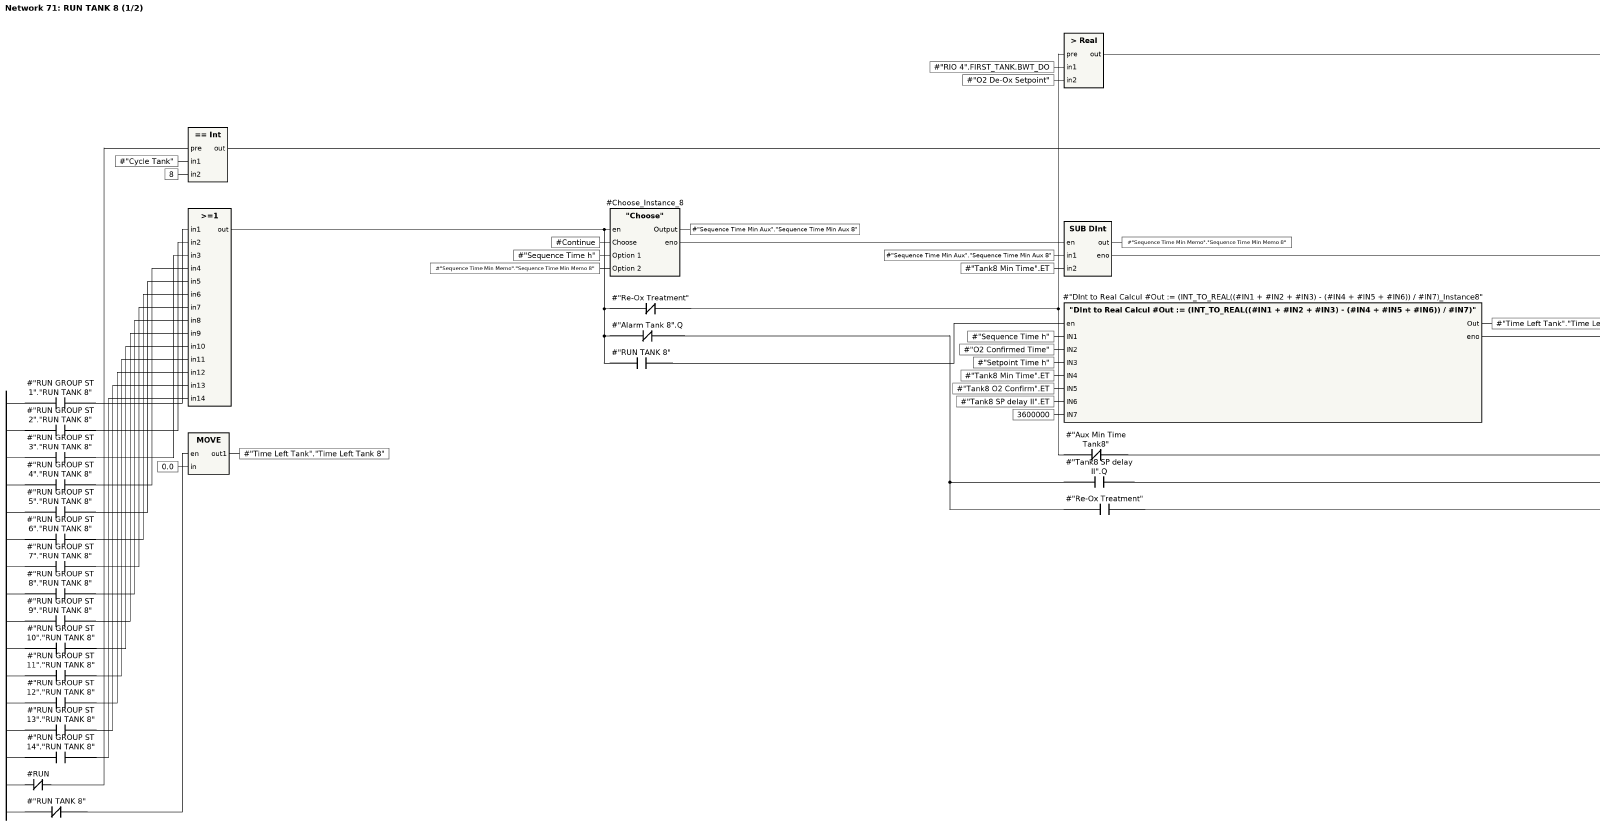
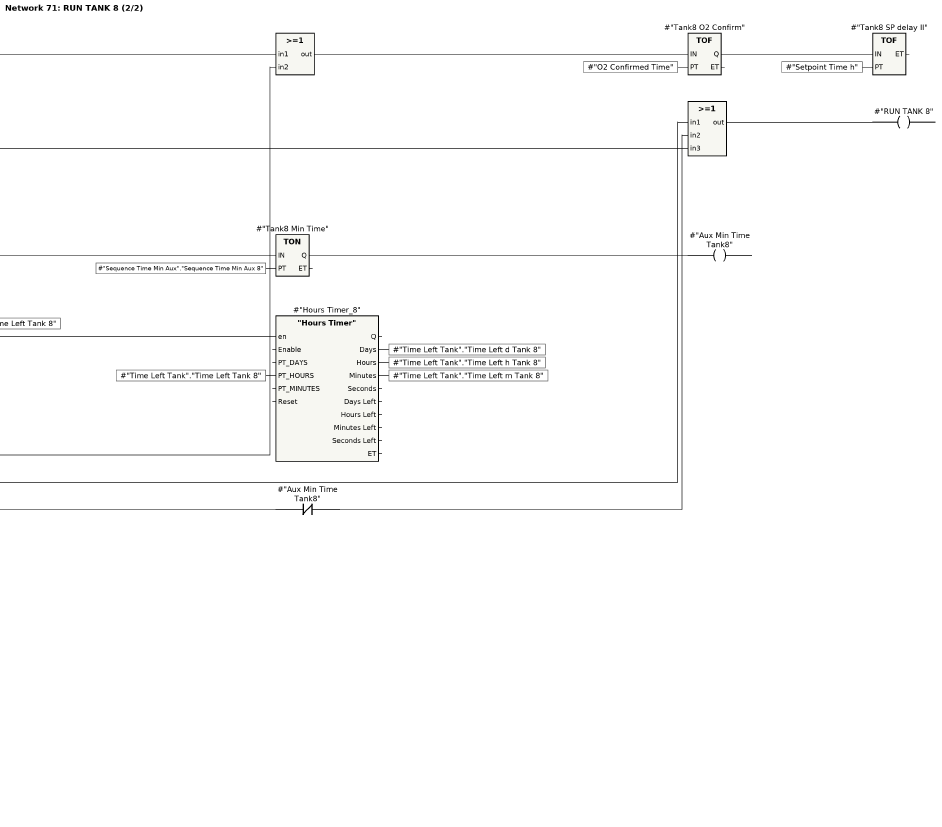
   #_w1 := #"RUN GROUP ST 1"."RUN TANK 8" OR #"RUN GROUP ST 2"."RUN TANK 8" OR #"RUN GROUP ST 3"."RUN TANK 8" OR #"RUN GROUP ST 4"."RUN TANK 8" OR #"RUN GROUP ST 5"."RUN TANK 8" OR #"RUN GROUP ST 6"."RUN TANK 8" OR #"RUN GROUP ST 7"."RUN TANK 8" OR #"RUN GROUP ST 8"."RUN TANK 8" OR #"RUN GROUP ST 9"."RUN TANK 8" OR #"RUN GROUP ST 10"."RUN TANK 8" OR #"RUN GROUP ST 11"."RUN TANK 8" OR #"RUN GROUP ST 12"."RUN TANK 8" OR #"RUN GROUP ST 13"."RUN TANK 8" OR #"RUN GROUP ST 14"."RUN TANK 8";
   #Choose_Instance_8(EN := #_w1,   // "Choose"
                      Choose := #Continue,
                      "Option 1" := #"Sequence Time h",
                      "Option 2" := #"Sequence Time Min Memo"."Sequence Time Min Memo 8",
                      Output => #"Sequence Time Min Aux"."Sequence Time Min Aux 8",
                      ENO => #_w2);
   IF #_w2 THEN
       #"Sequence Time Min Memo"."Sequence Time Min Memo 8" := #"Sequence Time Min Aux"."Sequence Time Min Aux 8" - #"Tank8 Min Time".ET;   // Memory of remained time for use to continue
   END_IF;
   #"Tank8 Min Time"(IN := #_w2, PT := #"Sequence Time Min Aux"."Sequence Time Min Aux 8");   // TON
   #"Aux Min Time Tank8" := #"Tank8 Min Time".Q;
   #"Tank8 O2 Confirm"(IN := #_w1 AND NOT #"Re-Ox Treatment" AND ((#"RIO 4".FIRST_TANK.BWT_DO > #"O2 De-Ox Setpoint") OR NOT #"Aux Min Time Tank8"),   // TOF
                       PT := #"O2 Confirmed Time");
   #"Tank8 SP delay II"(IN := #"Tank8 O2 Confirm".Q, PT := #"Setpoint Time h");   // TOF
   #"DInt to Real Calcul #Out := (INT_TO_REAL((#IN1 + #IN2 + #IN3) - (#IN4 + #IN5 + #IN6)) / #IN7)_Instance8"(EN := #_w1 AND #"RUN TANK 8",   // "DInt to Real Calcul #Out := (INT_TO_REAL((#IN1 + #IN2 + #IN3) - (#IN4 + #IN5 + #IN6)) / #IN7)"
                           IN1 := #"Sequence Time h",
                           IN2 := #"O2 Confirmed Time",
                           IN3 := #"Setpoint Time h",
                           IN4 := #"Tank8 Min Time".ET,
                           IN5 := #"Tank8 O2 Confirm".ET,
                           IN6 := #"Tank8 SP delay II".ET,
                           IN7 := 3600000,
                           Out => #"Time Left Tank"."Time Left Tank 8",
                           ENO => #_w3);
   IF #_w3 THEN
       #"Hours Timer_8"(PT_HOURS := #"Time Left Tank"."Time Left Tank 8",   // "Hours Timer"
                        Days => #"Time Left Tank"."Time Left d Tank 8",
                        Hours => #"Time Left Tank"."Time Left h Tank 8",
                        Minutes => #"Time Left Tank"."Time Left m Tank 8");
   END_IF;
   #"RUN TANK 8" := (#_w1 AND NOT #"Alarm Tank 8".Q AND (#"Tank8 SP delay II".Q OR (#"Re-Ox Treatment" AND NOT #"Aux Min Time Tank8"))) OR (NOT #RUN AND (#"Cycle Tank" = 8));
   IF NOT #"RUN TANK 8" THEN #"Time Left Tank"."Time Left Tank 8" := 0.0; END_IF;
END_REGION

REGION Network 72: RUN TANK 9
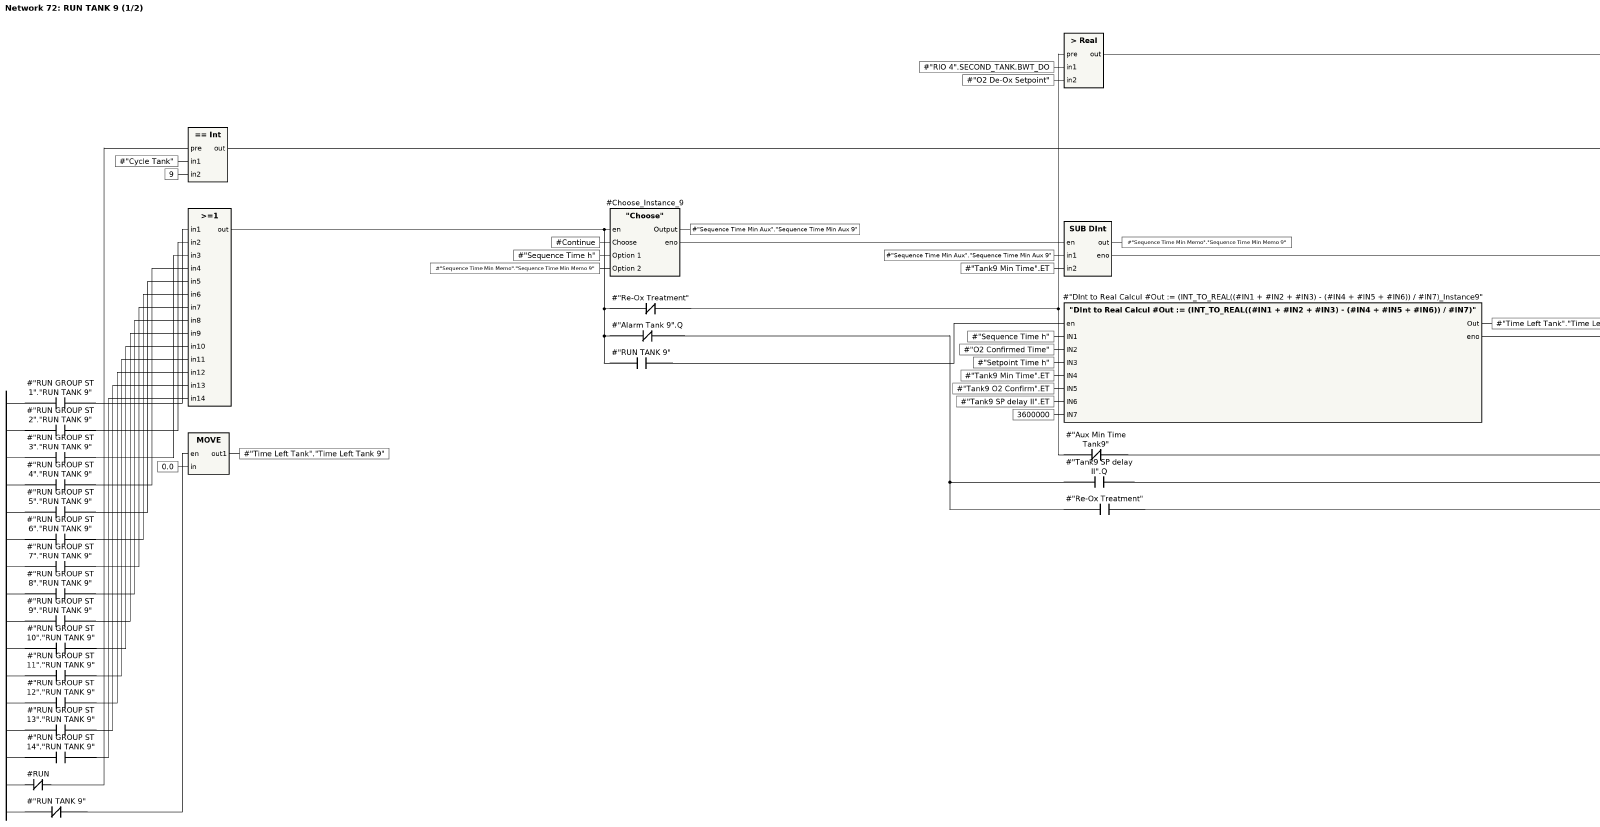
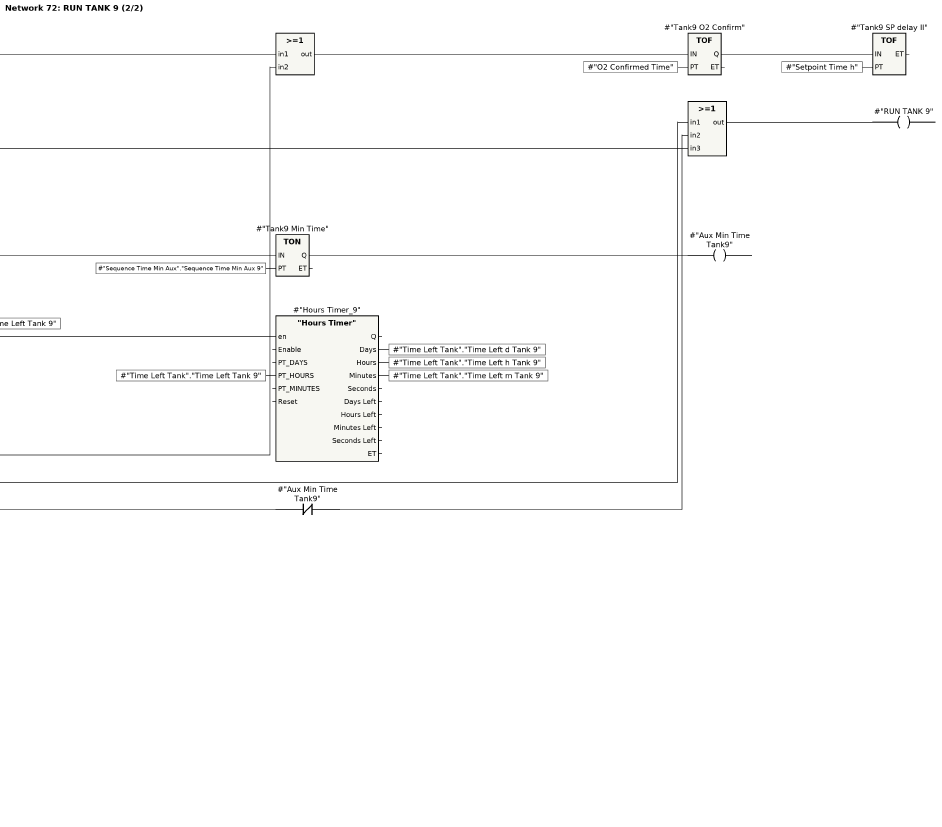
   #_w1 := #"RUN GROUP ST 1"."RUN TANK 9" OR #"RUN GROUP ST 2"."RUN TANK 9" OR #"RUN GROUP ST 3"."RUN TANK 9" OR #"RUN GROUP ST 4"."RUN TANK 9" OR #"RUN GROUP ST 5"."RUN TANK 9" OR #"RUN GROUP ST 6"."RUN TANK 9" OR #"RUN GROUP ST 7"."RUN TANK 9" OR #"RUN GROUP ST 8"."RUN TANK 9" OR #"RUN GROUP ST 9"."RUN TANK 9" OR #"RUN GROUP ST 10"."RUN TANK 9" OR #"RUN GROUP ST 11"."RUN TANK 9" OR #"RUN GROUP ST 12"."RUN TANK 9" OR #"RUN GROUP ST 13"."RUN TANK 9" OR #"RUN GROUP ST 14"."RUN TANK 9";
   #Choose_Instance_9(EN := #_w1,   // "Choose"
                      Choose := #Continue,
                      "Option 1" := #"Sequence Time h",
                      "Option 2" := #"Sequence Time Min Memo"."Sequence Time Min Memo 9",
                      Output => #"Sequence Time Min Aux"."Sequence Time Min Aux 9",
                      ENO => #_w2);
   IF #_w2 THEN
       #"Sequence Time Min Memo"."Sequence Time Min Memo 9" := #"Sequence Time Min Aux"."Sequence Time Min Aux 9" - #"Tank9 Min Time".ET;   // Memory of remained time for use to continue
   END_IF;
   #"Tank9 Min Time"(IN := #_w2, PT := #"Sequence Time Min Aux"."Sequence Time Min Aux 9");   // TON
   #"Aux Min Time Tank9" := #"Tank9 Min Time".Q;
   #"Tank9 O2 Confirm"(IN := #_w1 AND NOT #"Re-Ox Treatment" AND ((#"RIO 4".SECOND_TANK.BWT_DO > #"O2 De-Ox Setpoint") OR NOT #"Aux Min Time Tank9"),   // TOF
                       PT := #"O2 Confirmed Time");
   #"Tank9 SP delay II"(IN := #"Tank9 O2 Confirm".Q, PT := #"Setpoint Time h");   // TOF
   #"DInt to Real Calcul #Out := (INT_TO_REAL((#IN1 + #IN2 + #IN3) - (#IN4 + #IN5 + #IN6)) / #IN7)_Instance9"(EN := #_w1 AND #"RUN TANK 9",   // "DInt to Real Calcul #Out := (INT_TO_REAL((#IN1 + #IN2 + #IN3) - (#IN4 + #IN5 + #IN6)) / #IN7)"
                           IN1 := #"Sequence Time h",
                           IN2 := #"O2 Confirmed Time",
                           IN3 := #"Setpoint Time h",
                           IN4 := #"Tank9 Min Time".ET,
                           IN5 := #"Tank9 O2 Confirm".ET,
                           IN6 := #"Tank9 SP delay II".ET,
                           IN7 := 3600000,
                           Out => #"Time Left Tank"."Time Left Tank 9",
                           ENO => #_w3);
   IF #_w3 THEN
       #"Hours Timer_9"(PT_HOURS := #"Time Left Tank"."Time Left Tank 9",   // "Hours Timer"
                        Days => #"Time Left Tank"."Time Left d Tank 9",
                        Hours => #"Time Left Tank"."Time Left h Tank 9",
                        Minutes => #"Time Left Tank"."Time Left m Tank 9");
   END_IF;
   #"RUN TANK 9" := (#_w1 AND NOT #"Alarm Tank 9".Q AND (#"Tank9 SP delay II".Q OR (#"Re-Ox Treatment" AND NOT #"Aux Min Time Tank9"))) OR (NOT #RUN AND (#"Cycle Tank" = 9));
   IF NOT #"RUN TANK 9" THEN #"Time Left Tank"."Time Left Tank 9" := 0.0; END_IF;
END_REGION

REGION Network 73: RUN TANK 10
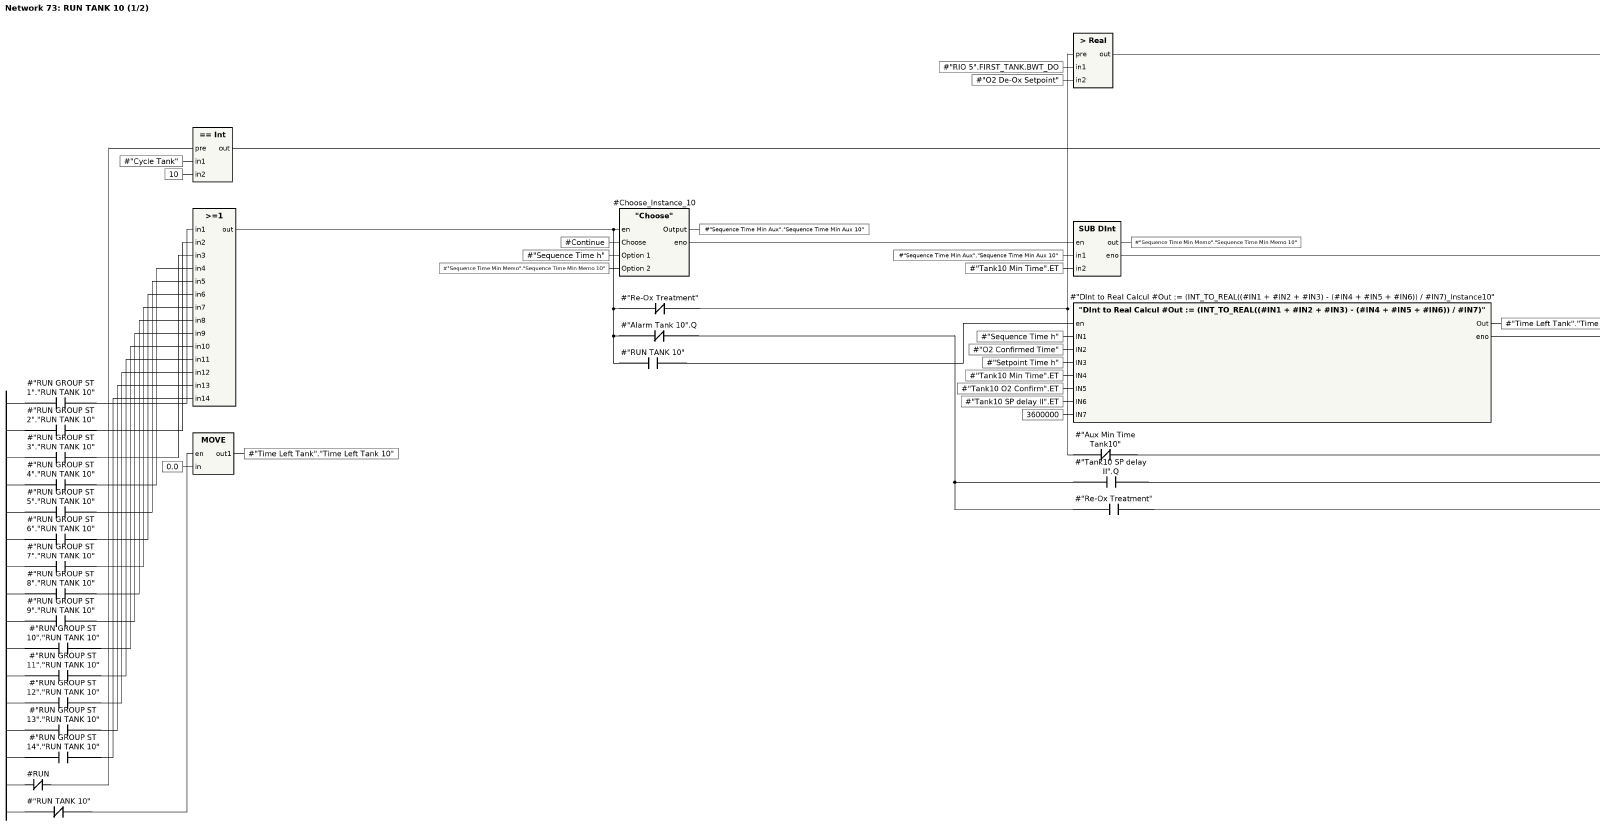
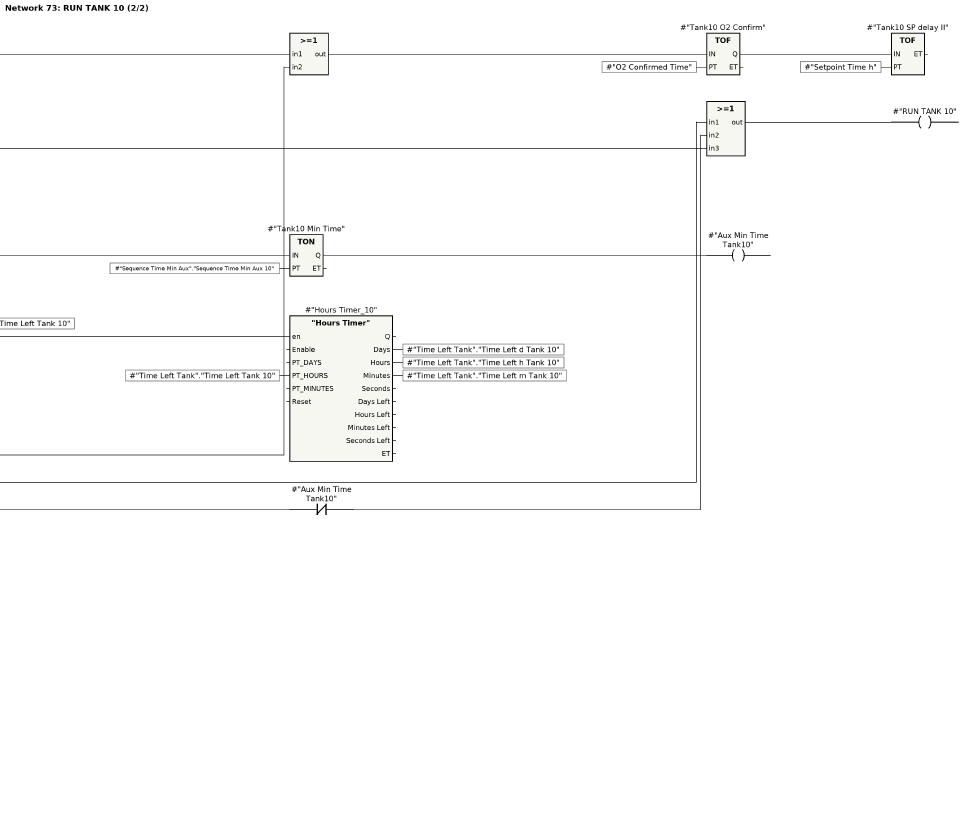
   #_w1 := #"RUN GROUP ST 1"."RUN TANK 10" OR #"RUN GROUP ST 2"."RUN TANK 10" OR #"RUN GROUP ST 3"."RUN TANK 10" OR #"RUN GROUP ST 4"."RUN TANK 10" OR #"RUN GROUP ST 5"."RUN TANK 10" OR #"RUN GROUP ST 6"."RUN TANK 10" OR #"RUN GROUP ST 7"."RUN TANK 10" OR #"RUN GROUP ST 8"."RUN TANK 10" OR #"RUN GROUP ST 9"."RUN TANK 10" OR #"RUN GROUP ST 10"."RUN TANK 10" OR #"RUN GROUP ST 11"."RUN TANK 10" OR #"RUN GROUP ST 12"."RUN TANK 10" OR #"RUN GROUP ST 13"."RUN TANK 10" OR #"RUN GROUP ST 14"."RUN TANK 10";
   #Choose_Instance_10(EN := #_w1,   // "Choose"
                       Choose := #Continue,
                       "Option 1" := #"Sequence Time h",
                       "Option 2" := #"Sequence Time Min Memo"."Sequence Time Min Memo 10",
                       Output => #"Sequence Time Min Aux"."Sequence Time Min Aux 10",
                       ENO => #_w2);
   IF #_w2 THEN
       #"Sequence Time Min Memo"."Sequence Time Min Memo 10" := #"Sequence Time Min Aux"."Sequence Time Min Aux 10" - #"Tank10 Min Time".ET;   // Memory of remained time for use to continue
   END_IF;
   #"Tank10 Min Time"(IN := #_w2, PT := #"Sequence Time Min Aux"."Sequence Time Min Aux 10");   // TON
   #"Aux Min Time Tank10" := #"Tank10 Min Time".Q;
   #"Tank10 O2 Confirm"(IN := #_w1 AND NOT #"Re-Ox Treatment" AND ((#"RIO 5".FIRST_TANK.BWT_DO > #"O2 De-Ox Setpoint") OR NOT #"Aux Min Time Tank10"),   // TOF
                        PT := #"O2 Confirmed Time");
   #"Tank10 SP delay II"(IN := #"Tank10 O2 Confirm".Q, PT := #"Setpoint Time h");   // TOF
   #"DInt to Real Calcul #Out := (INT_TO_REAL((#IN1 + #IN2 + #IN3) - (#IN4 + #IN5 + #IN6)) / #IN7)_Instance10"(EN := #_w1 AND #"RUN TANK 10",   // "DInt to Real Calcul #Out := (INT_TO_REAL((#IN1 + #IN2 + #IN3) - (#IN4 + #IN5 + #IN6)) / #IN7)"
                           IN1 := #"Sequence Time h",
                           IN2 := #"O2 Confirmed Time",
                           IN3 := #"Setpoint Time h",
                           IN4 := #"Tank10 Min Time".ET,
                           IN5 := #"Tank10 O2 Confirm".ET,
                           IN6 := #"Tank10 SP delay II".ET,
                           IN7 := 3600000,
                           Out => #"Time Left Tank"."Time Left Tank 10",
                           ENO => #_w3);
   IF #_w3 THEN
       #"Hours Timer_10"(PT_HOURS := #"Time Left Tank"."Time Left Tank 10",   // "Hours Timer"
                         Days => #"Time Left Tank"."Time Left d Tank 10",
                         Hours => #"Time Left Tank"."Time Left h Tank 10",
                         Minutes => #"Time Left Tank"."Time Left m Tank 10");
   END_IF;
   #"RUN TANK 10" := (#_w1 AND NOT #"Alarm Tank 10".Q AND (#"Tank10 SP delay II".Q OR (#"Re-Ox Treatment" AND NOT #"Aux Min Time Tank10"))) OR (NOT #RUN AND (#"Cycle Tank" = 10));
   IF NOT #"RUN TANK 10" THEN #"Time Left Tank"."Time Left Tank 10" := 0.0; END_IF;
END_REGION

REGION Network 74: RUN TANK 11
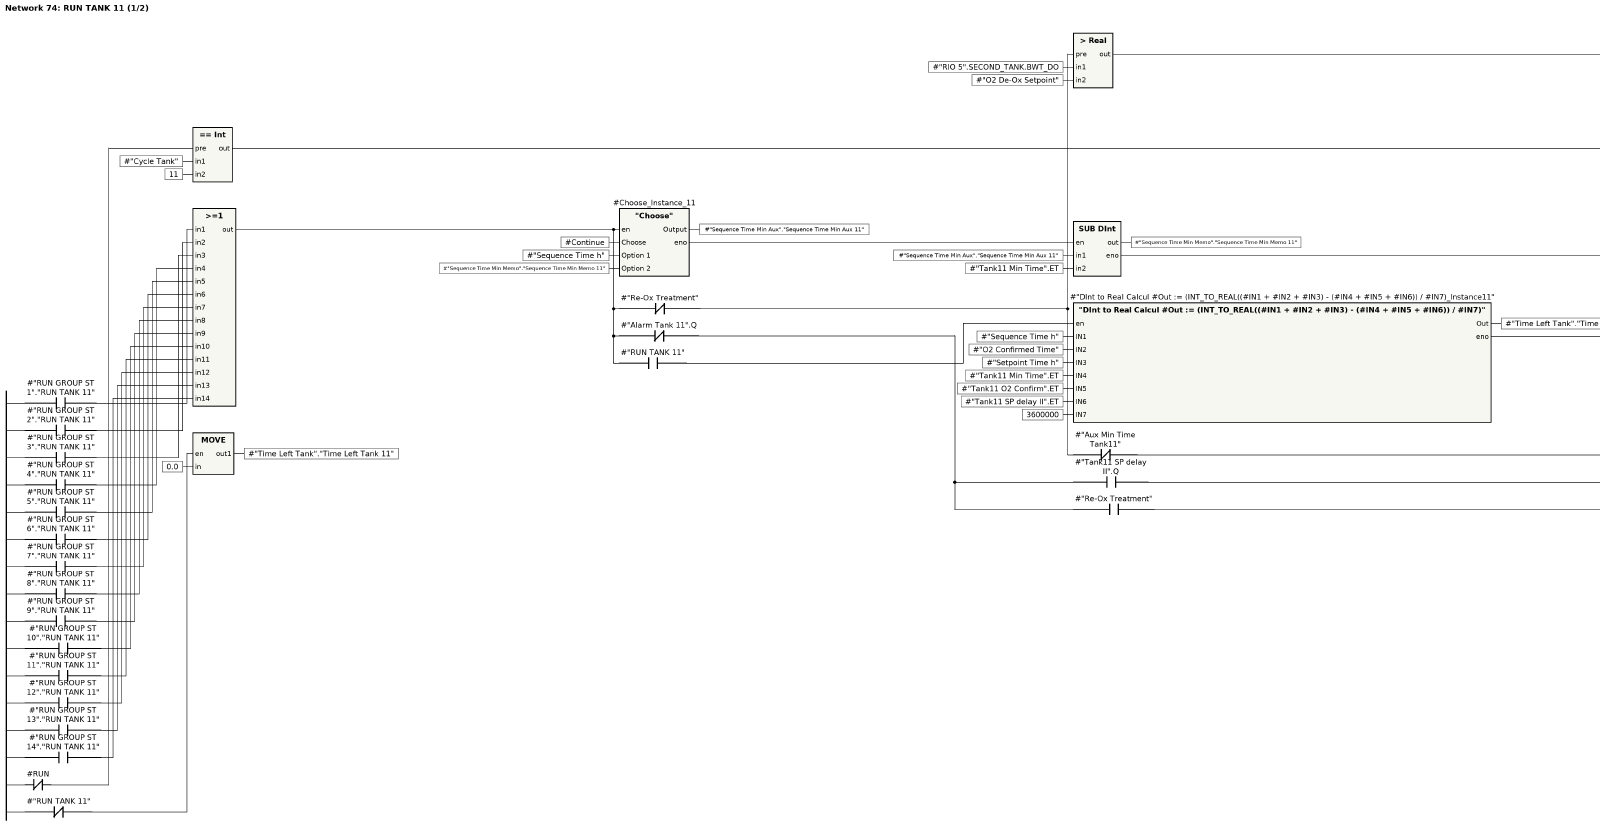
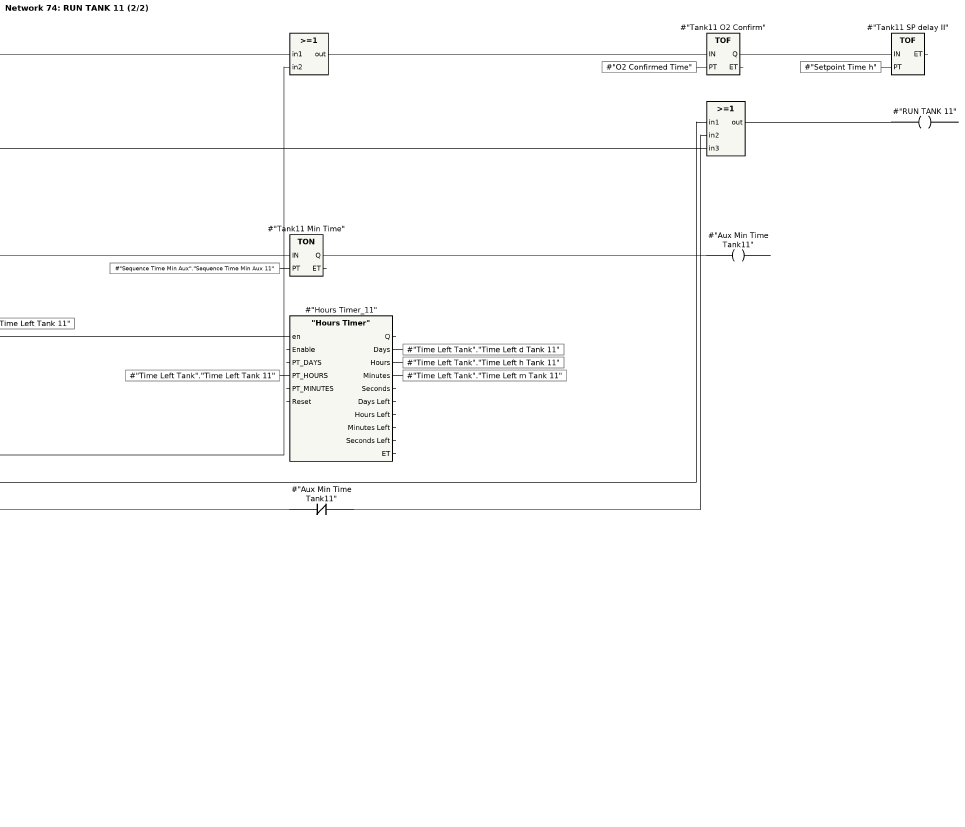
   #_w1 := #"RUN GROUP ST 1"."RUN TANK 11" OR #"RUN GROUP ST 2"."RUN TANK 11" OR #"RUN GROUP ST 3"."RUN TANK 11" OR #"RUN GROUP ST 4"."RUN TANK 11" OR #"RUN GROUP ST 5"."RUN TANK 11" OR #"RUN GROUP ST 6"."RUN TANK 11" OR #"RUN GROUP ST 7"."RUN TANK 11" OR #"RUN GROUP ST 8"."RUN TANK 11" OR #"RUN GROUP ST 9"."RUN TANK 11" OR #"RUN GROUP ST 10"."RUN TANK 11" OR #"RUN GROUP ST 11"."RUN TANK 11" OR #"RUN GROUP ST 12"."RUN TANK 11" OR #"RUN GROUP ST 13"."RUN TANK 11" OR #"RUN GROUP ST 14"."RUN TANK 11";
   #Choose_Instance_11(EN := #_w1,   // "Choose"
                       Choose := #Continue,
                       "Option 1" := #"Sequence Time h",
                       "Option 2" := #"Sequence Time Min Memo"."Sequence Time Min Memo 11",
                       Output => #"Sequence Time Min Aux"."Sequence Time Min Aux 11",
                       ENO => #_w2);
   IF #_w2 THEN
       #"Sequence Time Min Memo"."Sequence Time Min Memo 11" := #"Sequence Time Min Aux"."Sequence Time Min Aux 11" - #"Tank11 Min Time".ET;   // Memory of remained time for use to continue
   END_IF;
   #"Tank11 Min Time"(IN := #_w2, PT := #"Sequence Time Min Aux"."Sequence Time Min Aux 11");   // TON
   #"Aux Min Time Tank11" := #"Tank11 Min Time".Q;
   #"Tank11 O2 Confirm"(IN := #_w1 AND NOT #"Re-Ox Treatment" AND ((#"RIO 5".SECOND_TANK.BWT_DO > #"O2 De-Ox Setpoint") OR NOT #"Aux Min Time Tank11"),   // TOF
                        PT := #"O2 Confirmed Time");
   #"Tank11 SP delay II"(IN := #"Tank11 O2 Confirm".Q, PT := #"Setpoint Time h");   // TOF
   #"DInt to Real Calcul #Out := (INT_TO_REAL((#IN1 + #IN2 + #IN3) - (#IN4 + #IN5 + #IN6)) / #IN7)_Instance11"(EN := #_w1 AND #"RUN TANK 11",   // "DInt to Real Calcul #Out := (INT_TO_REAL((#IN1 + #IN2 + #IN3) - (#IN4 + #IN5 + #IN6)) / #IN7)"
                           IN1 := #"Sequence Time h",
                           IN2 := #"O2 Confirmed Time",
                           IN3 := #"Setpoint Time h",
                           IN4 := #"Tank11 Min Time".ET,
                           IN5 := #"Tank11 O2 Confirm".ET,
                           IN6 := #"Tank11 SP delay II".ET,
                           IN7 := 3600000,
                           Out => #"Time Left Tank"."Time Left Tank 11",
                           ENO => #_w3);
   IF #_w3 THEN
       #"Hours Timer_11"(PT_HOURS := #"Time Left Tank"."Time Left Tank 11",   // "Hours Timer"
                         Days => #"Time Left Tank"."Time Left d Tank 11",
                         Hours => #"Time Left Tank"."Time Left h Tank 11",
                         Minutes => #"Time Left Tank"."Time Left m Tank 11");
   END_IF;
   #"RUN TANK 11" := (#_w1 AND NOT #"Alarm Tank 11".Q AND (#"Tank11 SP delay II".Q OR (#"Re-Ox Treatment" AND NOT #"Aux Min Time Tank11"))) OR (NOT #RUN AND (#"Cycle Tank" = 11));
   IF NOT #"RUN TANK 11" THEN #"Time Left Tank"."Time Left Tank 11" := 0.0; END_IF;
END_REGION

REGION Network 75: RUN TANK 12
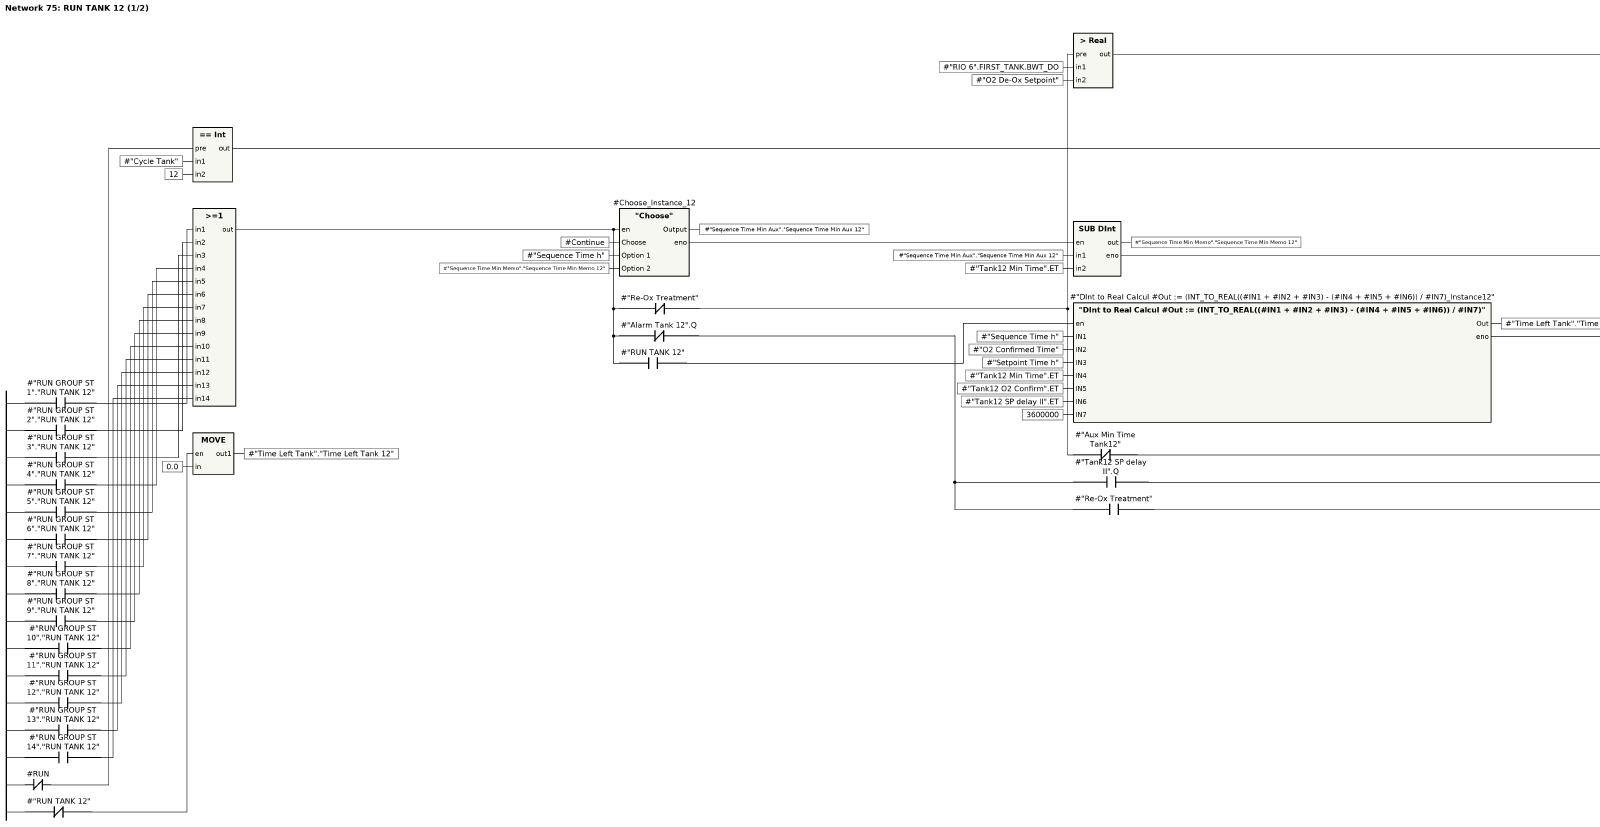
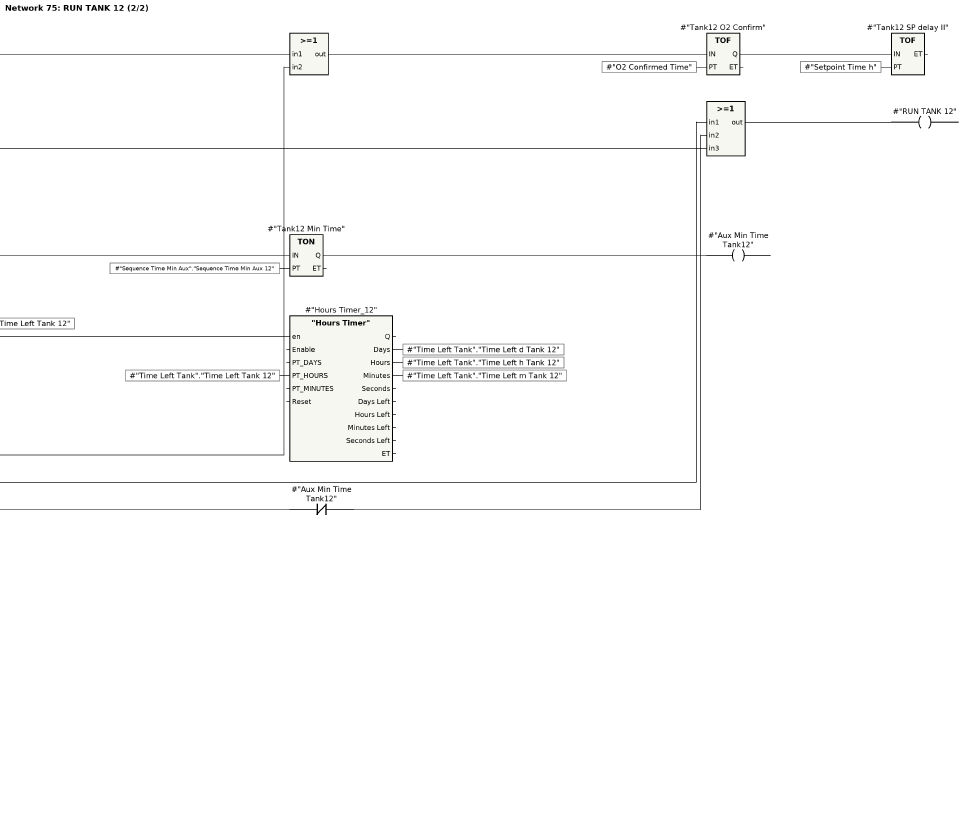
   #_w1 := #"RUN GROUP ST 1"."RUN TANK 12" OR #"RUN GROUP ST 2"."RUN TANK 12" OR #"RUN GROUP ST 3"."RUN TANK 12" OR #"RUN GROUP ST 4"."RUN TANK 12" OR #"RUN GROUP ST 5"."RUN TANK 12" OR #"RUN GROUP ST 6"."RUN TANK 12" OR #"RUN GROUP ST 7"."RUN TANK 12" OR #"RUN GROUP ST 8"."RUN TANK 12" OR #"RUN GROUP ST 9"."RUN TANK 12" OR #"RUN GROUP ST 10"."RUN TANK 12" OR #"RUN GROUP ST 11"."RUN TANK 12" OR #"RUN GROUP ST 12"."RUN TANK 12" OR #"RUN GROUP ST 13"."RUN TANK 12" OR #"RUN GROUP ST 14"."RUN TANK 12";
   #Choose_Instance_12(EN := #_w1,   // "Choose"
                       Choose := #Continue,
                       "Option 1" := #"Sequence Time h",
                       "Option 2" := #"Sequence Time Min Memo"."Sequence Time Min Memo 12",
                       Output => #"Sequence Time Min Aux"."Sequence Time Min Aux 12",
                       ENO => #_w2);
   IF #_w2 THEN
       #"Sequence Time Min Memo"."Sequence Time Min Memo 12" := #"Sequence Time Min Aux"."Sequence Time Min Aux 12" - #"Tank12 Min Time".ET;   // Memory of remained time for use to continue
   END_IF;
   #"Tank12 Min Time"(IN := #_w2, PT := #"Sequence Time Min Aux"."Sequence Time Min Aux 12");   // TON
   #"Aux Min Time Tank12" := #"Tank12 Min Time".Q;
   #"Tank12 O2 Confirm"(IN := #_w1 AND NOT #"Re-Ox Treatment" AND ((#"RIO 6".FIRST_TANK.BWT_DO > #"O2 De-Ox Setpoint") OR NOT #"Aux Min Time Tank12"),   // TOF
                        PT := #"O2 Confirmed Time");
   #"Tank12 SP delay II"(IN := #"Tank12 O2 Confirm".Q, PT := #"Setpoint Time h");   // TOF
   #"DInt to Real Calcul #Out := (INT_TO_REAL((#IN1 + #IN2 + #IN3) - (#IN4 + #IN5 + #IN6)) / #IN7)_Instance12"(EN := #_w1 AND #"RUN TANK 12",   // "DInt to Real Calcul #Out := (INT_TO_REAL((#IN1 + #IN2 + #IN3) - (#IN4 + #IN5 + #IN6)) / #IN7)"
                           IN1 := #"Sequence Time h",
                           IN2 := #"O2 Confirmed Time",
                           IN3 := #"Setpoint Time h",
                           IN4 := #"Tank12 Min Time".ET,
                           IN5 := #"Tank12 O2 Confirm".ET,
                           IN6 := #"Tank12 SP delay II".ET,
                           IN7 := 3600000,
                           Out => #"Time Left Tank"."Time Left Tank 12",
                           ENO => #_w3);
   IF #_w3 THEN
       #"Hours Timer_12"(PT_HOURS := #"Time Left Tank"."Time Left Tank 12",   // "Hours Timer"
                         Days => #"Time Left Tank"."Time Left d Tank 12",
                         Hours => #"Time Left Tank"."Time Left h Tank 12",
                         Minutes => #"Time Left Tank"."Time Left m Tank 12");
   END_IF;
   #"RUN TANK 12" := (#_w1 AND NOT #"Alarm Tank 12".Q AND (#"Tank12 SP delay II".Q OR (#"Re-Ox Treatment" AND NOT #"Aux Min Time Tank12"))) OR (NOT #RUN AND (#"Cycle Tank" = 12));
   IF NOT #"RUN TANK 12" THEN #"Time Left Tank"."Time Left Tank 12" := 0.0; END_IF;
END_REGION

REGION Network 76: RUN TANK 13
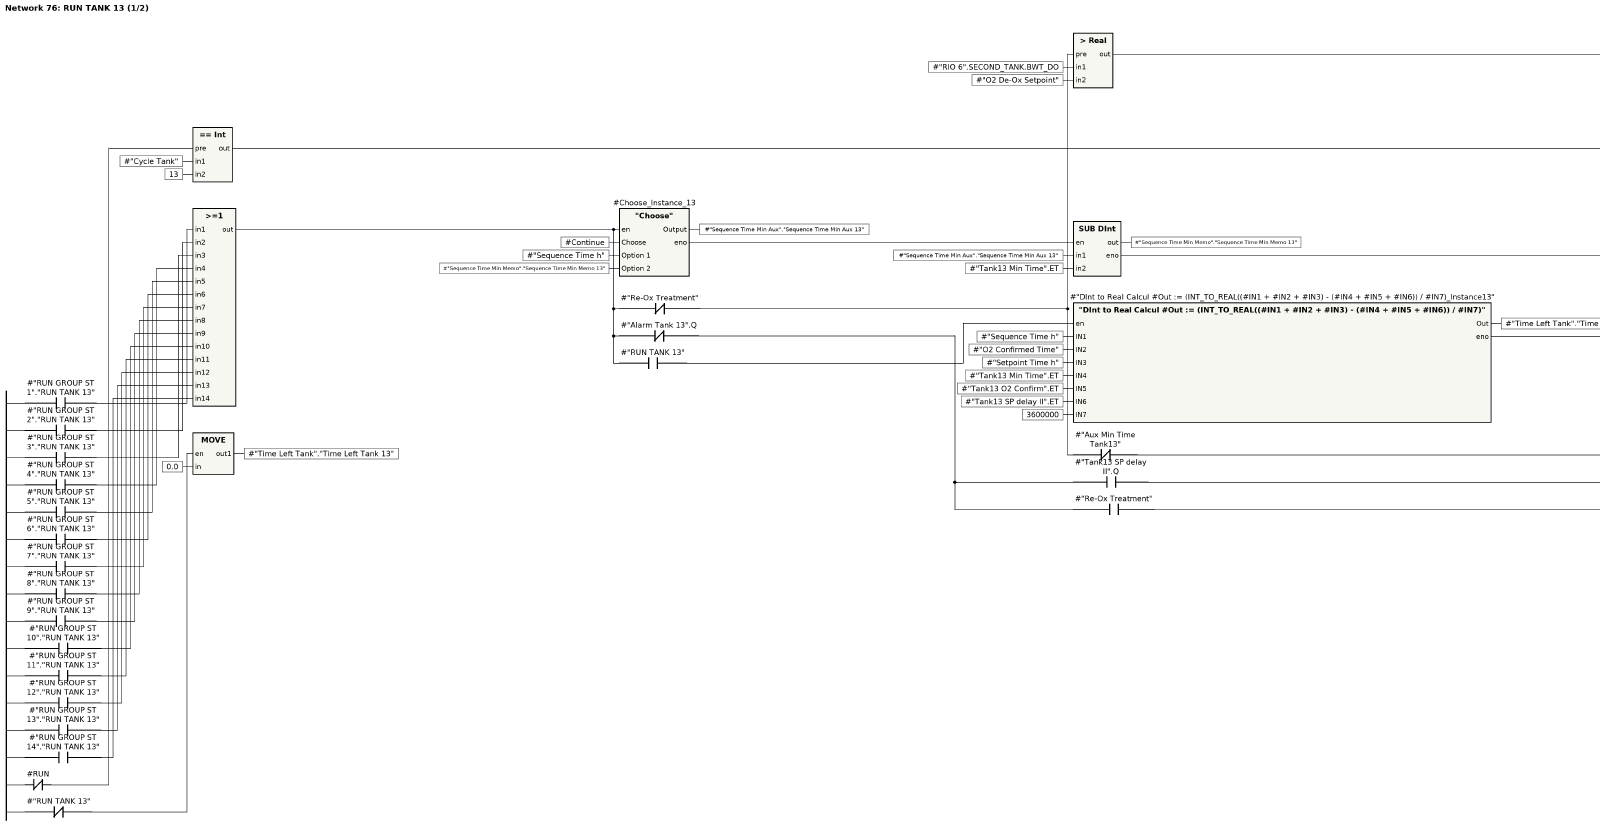
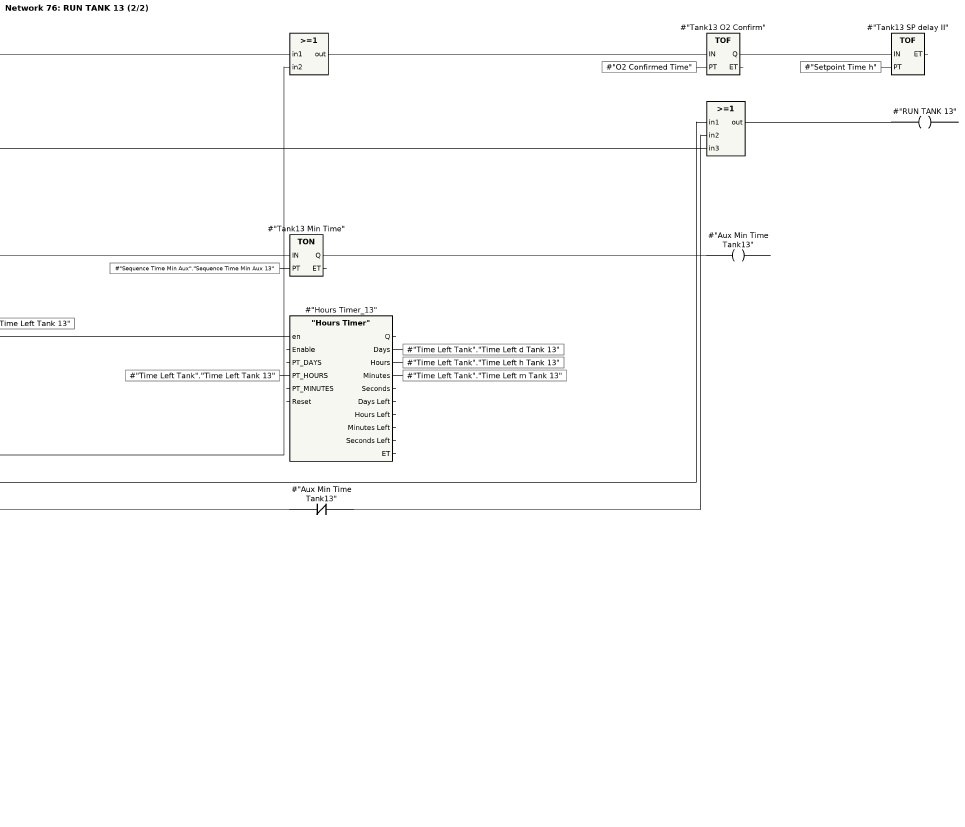
   #_w1 := #"RUN GROUP ST 1"."RUN TANK 13" OR #"RUN GROUP ST 2"."RUN TANK 13" OR #"RUN GROUP ST 3"."RUN TANK 13" OR #"RUN GROUP ST 4"."RUN TANK 13" OR #"RUN GROUP ST 5"."RUN TANK 13" OR #"RUN GROUP ST 6"."RUN TANK 13" OR #"RUN GROUP ST 7"."RUN TANK 13" OR #"RUN GROUP ST 8"."RUN TANK 13" OR #"RUN GROUP ST 9"."RUN TANK 13" OR #"RUN GROUP ST 10"."RUN TANK 13" OR #"RUN GROUP ST 11"."RUN TANK 13" OR #"RUN GROUP ST 12"."RUN TANK 13" OR #"RUN GROUP ST 13"."RUN TANK 13" OR #"RUN GROUP ST 14"."RUN TANK 13";
   #Choose_Instance_13(EN := #_w1,   // "Choose"
                       Choose := #Continue,
                       "Option 1" := #"Sequence Time h",
                       "Option 2" := #"Sequence Time Min Memo"."Sequence Time Min Memo 13",
                       Output => #"Sequence Time Min Aux"."Sequence Time Min Aux 13",
                       ENO => #_w2);
   IF #_w2 THEN
       #"Sequence Time Min Memo"."Sequence Time Min Memo 13" := #"Sequence Time Min Aux"."Sequence Time Min Aux 13" - #"Tank13 Min Time".ET;   // Memory of remained time for use to continue
   END_IF;
   #"Tank13 Min Time"(IN := #_w2, PT := #"Sequence Time Min Aux"."Sequence Time Min Aux 13");   // TON
   #"Aux Min Time Tank13" := #"Tank13 Min Time".Q;
   #"Tank13 O2 Confirm"(IN := #_w1 AND NOT #"Re-Ox Treatment" AND ((#"RIO 6".SECOND_TANK.BWT_DO > #"O2 De-Ox Setpoint") OR NOT #"Aux Min Time Tank13"),   // TOF
                        PT := #"O2 Confirmed Time");
   #"Tank13 SP delay II"(IN := #"Tank13 O2 Confirm".Q, PT := #"Setpoint Time h");   // TOF
   #"DInt to Real Calcul #Out := (INT_TO_REAL((#IN1 + #IN2 + #IN3) - (#IN4 + #IN5 + #IN6)) / #IN7)_Instance13"(EN := #_w1 AND #"RUN TANK 13",   // "DInt to Real Calcul #Out := (INT_TO_REAL((#IN1 + #IN2 + #IN3) - (#IN4 + #IN5 + #IN6)) / #IN7)"
                           IN1 := #"Sequence Time h",
                           IN2 := #"O2 Confirmed Time",
                           IN3 := #"Setpoint Time h",
                           IN4 := #"Tank13 Min Time".ET,
                           IN5 := #"Tank13 O2 Confirm".ET,
                           IN6 := #"Tank13 SP delay II".ET,
                           IN7 := 3600000,
                           Out => #"Time Left Tank"."Time Left Tank 13",
                           ENO => #_w3);
   IF #_w3 THEN
       #"Hours Timer_13"(PT_HOURS := #"Time Left Tank"."Time Left Tank 13",   // "Hours Timer"
                         Days => #"Time Left Tank"."Time Left d Tank 13",
                         Hours => #"Time Left Tank"."Time Left h Tank 13",
                         Minutes => #"Time Left Tank"."Time Left m Tank 13");
   END_IF;
   #"RUN TANK 13" := (#_w1 AND NOT #"Alarm Tank 13".Q AND (#"Tank13 SP delay II".Q OR (#"Re-Ox Treatment" AND NOT #"Aux Min Time Tank13"))) OR (NOT #RUN AND (#"Cycle Tank" = 13));
   IF NOT #"RUN TANK 13" THEN #"Time Left Tank"."Time Left Tank 13" := 0.0; END_IF;
END_REGION

REGION Network 77: RUN TANK 14
